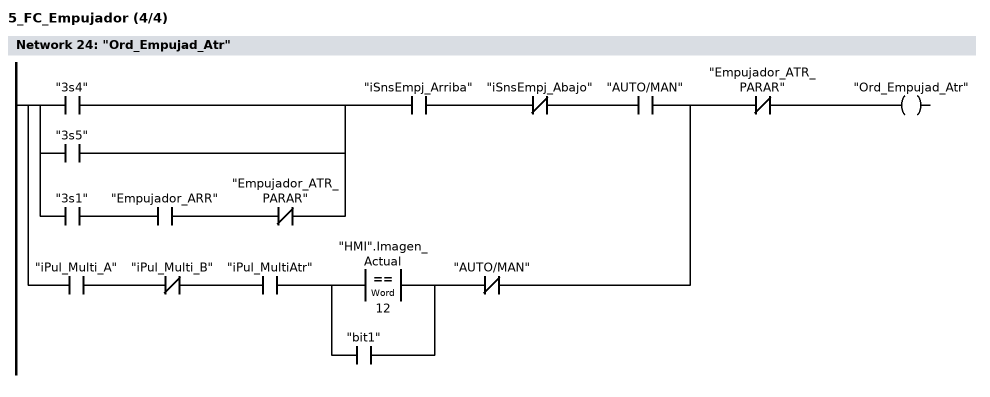
   RUNG wire#powerrail
      Contact( "3s4" )
      wire#w1
      Contact( "iSnsEmpj_Arriba" )
      I_Contact( "iSnsEmpj_Abajo" )
      Contact( "AUTO/MAN" )
      wire#w2
      I_Contact( "Empujador_ATR_PARAR" )
      Coil( "Ord_Empujad_Atr" )
   END_RUNG
   RUNG wire#powerrail
      Contact( "3s5" )
   END_RUNG wire#w1
   RUNG wire#powerrail
      Contact( "3s1" )
      Contact( "Empujador_ARR" )
      I_Contact( "Empujador_ATR_PARAR" )
   END_RUNG wire#w1
   RUNG wire#powerrail
      Contact( "iPul_Multi_A" )
      I_Contact( "iPul_Multi_B" )
      Contact( "iPul_MultiAtr" )
      wire#w3
      { S7_Templates := "SrcType := Word" } EQ_Contact(in1 := "HMI".Imagen_Actual, in2 := 12)
      wire#w4
      I_Contact( "AUTO/MAN" )
   END_RUNG wire#w2
   RUNG wire#w3
      Contact( "bit1" )
   END_RUNG wire#w4
   // the same network as SCL:
   "Ord_Empujad_Atr" := ((("3s4" OR "3s5" OR ("3s1" AND "Empujador_ARR" AND NOT "Empujador_ATR_PARAR")) AND "iSnsEmpj_Arriba" AND NOT "iSnsEmpj_Abajo" AND "AUTO/MAN") OR ("iPul_Multi_A" AND NOT "iPul_Multi_B" AND "iPul_MultiAtr" AND (("HMI".Imagen_Actual = 12) OR "bit1") AND NOT "AUTO/MAN")) AND NOT "Empujador_ATR_PARAR";
END_REGION
END_FUNCTION

FUNCTION "6_FC_Carga_Pallets" : Void   // FC13, LAD
{ S7_Optimized_Access := 'FALSE' }
VERSION : 0.1
BEGIN

REGION Network 1: "Poner_Mordazas"
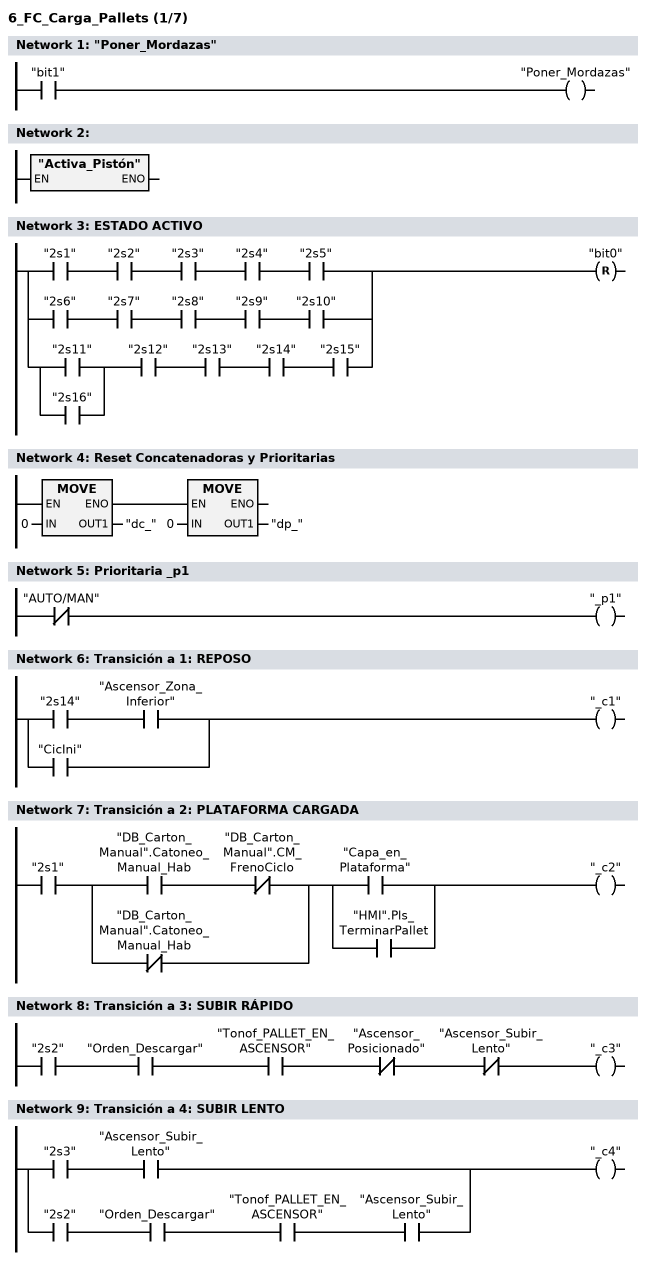
   RUNG wire#powerrail
      Contact( "bit1" )
      Coil( "Poner_Mordazas" )
   END_RUNG
   // the same network as SCL:
   "Poner_Mordazas" := "bit1";
END_REGION

REGION Network 2
   RUNG wire#powerrail
      "Activa_Pistón"()
   END_RUNG
   // the same network as SCL:
   "Activa_Pistón"();
END_REGION

REGION Network 3: ESTADO ACTIVO
   RUNG wire#powerrail
      Contact( "2s1" )
      Contact( "2s2" )
      Contact( "2s3" )
      Contact( "2s4" )
      Contact( "2s5" )
      wire#w1
      R_Coil( "bit0" )
   END_RUNG
   RUNG wire#powerrail
      Contact( "2s6" )
      Contact( "2s7" )
      Contact( "2s8" )
      Contact( "2s9" )
      Contact( "2s10" )
   END_RUNG wire#w1
   RUNG wire#powerrail
      Contact( "2s11" )
      wire#w2
      Contact( "2s12" )
      Contact( "2s13" )
      Contact( "2s14" )
      Contact( "2s15" )
   END_RUNG wire#w1
   RUNG wire#powerrail
      Contact( "2s16" )
   END_RUNG wire#w2
   // the same network as SCL:
   IF ("2s1" AND "2s2" AND "2s3" AND "2s4" AND "2s5") OR ("2s6" AND "2s7" AND "2s8" AND "2s9" AND "2s10") OR (("2s11" OR "2s16") AND "2s12" AND "2s13" AND "2s14" AND "2s15") THEN
       "bit0" := FALSE;
   END_IF;
END_REGION

REGION Network 4: Reset Concatenadoras y Prioritarias
   RUNG wire#powerrail
      { S7_GenerateENO := "TRUE" } Move(in := 0, out1 => "dc_")
      { S7_GenerateENO := "TRUE" } Move(in := 0, out1 => "dp_")
   END_RUNG
   // the same network as SCL:
   // ENO of a box is taken as its EN; it also drops when the box reports an error
   "dc_" := 0;
   "dp_" := 0;
END_REGION

REGION Network 5: Prioritaria _p1
   RUNG wire#powerrail
      I_Contact( "AUTO/MAN" )
      Coil( "_p1" )
   END_RUNG
   // the same network as SCL:
   "_p1" := NOT "AUTO/MAN";
END_REGION

REGION Network 6: Transición a 1: REPOSO
   RUNG wire#powerrail
      Contact( "2s14" )
      Contact( "Ascensor_Zona_Inferior" )
      wire#w1
      Coil( "_c1" )
   END_RUNG
   RUNG wire#powerrail
      Contact( "CicIni" )
   END_RUNG wire#w1
   // the same network as SCL:
   "_c1" := ("2s14" AND "Ascensor_Zona_Inferior") OR "CicIni";
END_REGION

REGION Network 7: Transición a 2: PLATAFORMA CARGADA
   RUNG wire#powerrail
      Contact( "2s1" )
      wire#w1
      Contact( "DB_Carton_Manual".Catoneo_Manual_Hab )
      I_Contact( "DB_Carton_Manual".CM_FrenoCiclo )
      wire#w2
      Contact( "Capa_en_Plataforma" )
      wire#w3
      Coil( "_c2" )
   END_RUNG
   RUNG wire#w1
      I_Contact( "DB_Carton_Manual".Catoneo_Manual_Hab )
   END_RUNG wire#w2
   RUNG wire#w2
      Contact( "HMI".Pls_TerminarPallet )
   END_RUNG wire#w3
   // the same network as SCL:
   "_c2" := "2s1" AND (("DB_Carton_Manual".Catoneo_Manual_Hab AND NOT "DB_Carton_Manual".CM_FrenoCiclo) OR NOT "DB_Carton_Manual".Catoneo_Manual_Hab) AND ("Capa_en_Plataforma" OR "HMI".Pls_TerminarPallet);
END_REGION

REGION Network 8: Transición a 3: SUBIR RÁPIDO
   RUNG wire#powerrail
      Contact( "2s2" )
      Contact( "Orden_Descargar" )
      Contact( "Tonof_PALLET_EN_ASCENSOR" )
      I_Contact( "Ascensor_Posicionado" )
      I_Contact( "Ascensor_Subir_Lento" )
      Coil( "_c3" )
   END_RUNG
   // the same network as SCL:
   "_c3" := "2s2" AND "Orden_Descargar" AND "Tonof_PALLET_EN_ASCENSOR" AND NOT "Ascensor_Posicionado" AND NOT "Ascensor_Subir_Lento";
END_REGION

REGION Network 9: Transición a 4: SUBIR LENTO
   RUNG wire#powerrail
      Contact( "2s3" )
      Contact( "Ascensor_Subir_Lento" )
      wire#w1
      Coil( "_c4" )
   END_RUNG
   RUNG wire#powerrail
      Contact( "2s2" )
      Contact( "Orden_Descargar" )
      Contact( "Tonof_PALLET_EN_ASCENSOR" )
      Contact( "Ascensor_Subir_Lento" )
   END_RUNG wire#w1
   // the same network as SCL:
   "_c4" := ("2s3" AND "Ascensor_Subir_Lento") OR ("2s2" AND "Orden_Descargar" AND "Tonof_PALLET_EN_ASCENSOR" AND "Ascensor_Subir_Lento");
END_REGION

REGION Network 10: Transición a 5: ADELANTAR
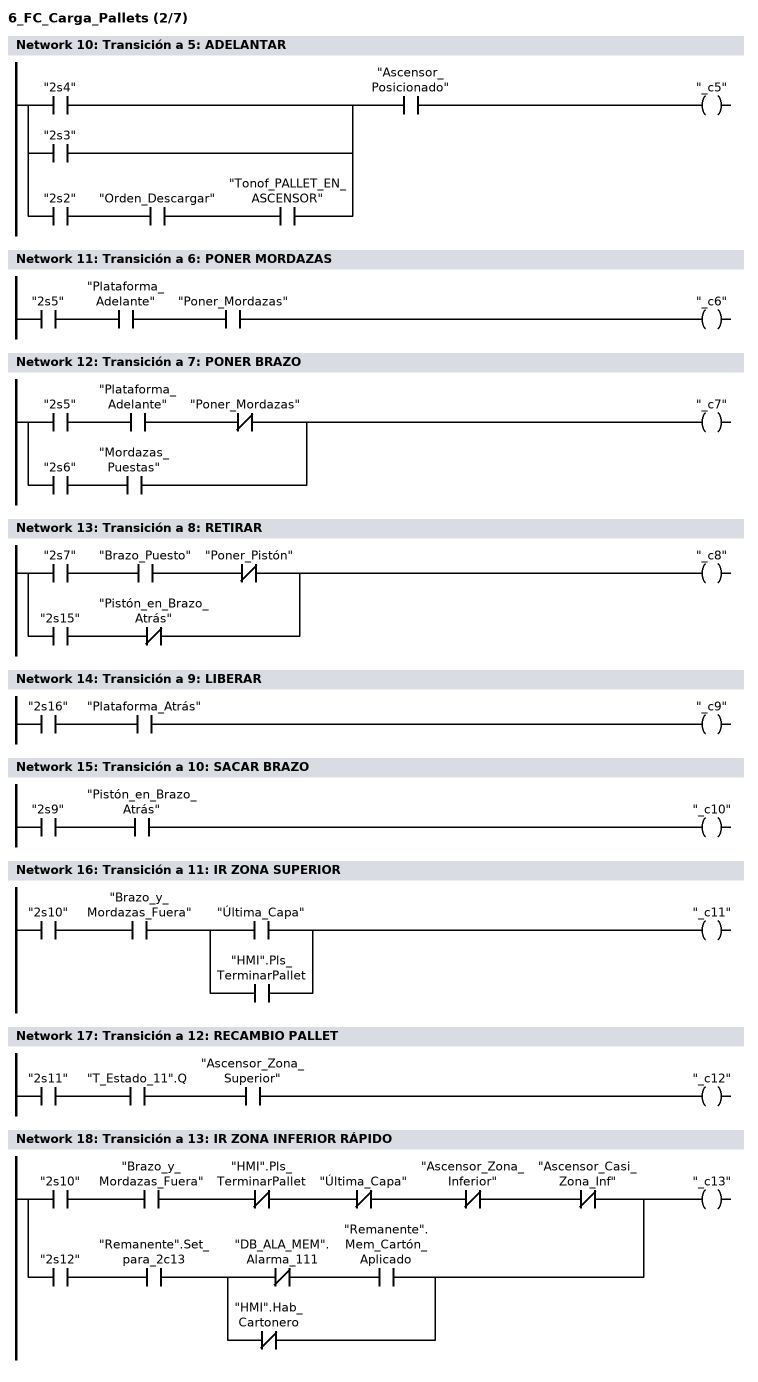
   RUNG wire#powerrail
      Contact( "2s4" )
      wire#w1
      Contact( "Ascensor_Posicionado" )
      Coil( "_c5" )
   END_RUNG
   RUNG wire#powerrail
      Contact( "2s3" )
   END_RUNG wire#w1
   RUNG wire#powerrail
      Contact( "2s2" )
      Contact( "Orden_Descargar" )
      Contact( "Tonof_PALLET_EN_ASCENSOR" )
   END_RUNG wire#w1
   // the same network as SCL:
   "_c5" := ("2s4" OR "2s3" OR ("2s2" AND "Orden_Descargar" AND "Tonof_PALLET_EN_ASCENSOR")) AND "Ascensor_Posicionado";
END_REGION

REGION Network 11: Transición a 6: PONER MORDAZAS
   RUNG wire#powerrail
      Contact( "2s5" )
      Contact( "Plataforma_Adelante" )
      Contact( "Poner_Mordazas" )
      Coil( "_c6" )
   END_RUNG
   // the same network as SCL:
   "_c6" := "2s5" AND "Plataforma_Adelante" AND "Poner_Mordazas";
END_REGION

REGION Network 12: Transición a 7: PONER BRAZO
   RUNG wire#powerrail
      Contact( "2s5" )
      Contact( "Plataforma_Adelante" )
      I_Contact( "Poner_Mordazas" )
      wire#w1
      Coil( "_c7" )
   END_RUNG
   RUNG wire#powerrail
      Contact( "2s6" )
      Contact( "Mordazas_Puestas" )
   END_RUNG wire#w1
   // the same network as SCL:
   "_c7" := ("2s5" AND "Plataforma_Adelante" AND NOT "Poner_Mordazas") OR ("2s6" AND "Mordazas_Puestas");
END_REGION

REGION Network 13: Transición a 8: RETIRAR
   RUNG wire#powerrail
      Contact( "2s7" )
      Contact( "Brazo_Puesto" )
      I_Contact( "Poner_Pistón" )
      wire#w1
      Coil( "_c8" )
   END_RUNG
   RUNG wire#powerrail
      Contact( "2s15" )
      I_Contact( "Pistón_en_Brazo_Atrás" )
   END_RUNG wire#w1
   // the same network as SCL:
   "_c8" := ("2s7" AND "Brazo_Puesto" AND NOT "Poner_Pistón") OR ("2s15" AND NOT "Pistón_en_Brazo_Atrás");
END_REGION

REGION Network 14: Transición a 9: LIBERAR
   RUNG wire#powerrail
      Contact( "2s16" )
      Contact( "Plataforma_Atrás" )
      Coil( "_c9" )
   END_RUNG
   // the same network as SCL:
   "_c9" := "2s16" AND "Plataforma_Atrás";
END_REGION

REGION Network 15: Transición a 10: SACAR BRAZO
   RUNG wire#powerrail
      Contact( "2s9" )
      Contact( "Pistón_en_Brazo_Atrás" )
      Coil( "_c10" )
   END_RUNG
   // the same network as SCL:
   "_c10" := "2s9" AND "Pistón_en_Brazo_Atrás";
END_REGION

REGION Network 16: Transición a 11: IR ZONA SUPERIOR
   RUNG wire#powerrail
      Contact( "2s10" )
      Contact( "Brazo_y_Mordazas_Fuera" )
      wire#w1
      Contact( "Última_Capa" )
      wire#w2
      Coil( "_c11" )
   END_RUNG
   RUNG wire#w1
      Contact( "HMI".Pls_TerminarPallet )
   END_RUNG wire#w2
   // the same network as SCL:
   "_c11" := "2s10" AND "Brazo_y_Mordazas_Fuera" AND ("Última_Capa" OR "HMI".Pls_TerminarPallet);
END_REGION

REGION Network 17: Transición a 12: RECAMBIO PALLET
   RUNG wire#powerrail
      Contact( "2s11" )
      Contact( "T_Estado_11".Q )
      Contact( "Ascensor_Zona_Superior" )
      Coil( "_c12" )
   END_RUNG
   // the same network as SCL:
   "_c12" := "2s11" AND "T_Estado_11".Q AND "Ascensor_Zona_Superior";
END_REGION

REGION Network 18: Transición a 13: IR ZONA INFERIOR RÁPIDO
   RUNG wire#powerrail
      Contact( "2s10" )
      Contact( "Brazo_y_Mordazas_Fuera" )
      I_Contact( "HMI".Pls_TerminarPallet )
      I_Contact( "Última_Capa" )
      I_Contact( "Ascensor_Zona_Inferior" )
      I_Contact( "Ascensor_Casi_Zona_Inf" )
      wire#w1
      Coil( "_c13" )
   END_RUNG
   RUNG wire#powerrail
      Contact( "2s12" )
      Contact( "Remanente".Set_para_2c13 )
      wire#w2
      I_Contact( "DB_ALA_MEM".Alarma_111 )
      Contact( "Remanente".Mem_Cartón_Aplicado )
   END_RUNG wire#w1
   RUNG wire#w2
      I_Contact( "HMI".Hab_Cartonero )
   END_RUNG wire#w1
   // the same network as SCL:
   "_c13" := ("2s10" AND "Brazo_y_Mordazas_Fuera" AND NOT "HMI".Pls_TerminarPallet AND NOT "Última_Capa" AND NOT "Ascensor_Zona_Inferior" AND NOT "Ascensor_Casi_Zona_Inf") OR ("2s12" AND "Remanente".Set_para_2c13 AND ((NOT "DB_ALA_MEM".Alarma_111 AND "Remanente".Mem_Cartón_Aplicado) OR NOT "HMI".Hab_Cartonero));
END_REGION

REGION Network 19: Transición a 14: IR ZONA INFERIOR LENTO
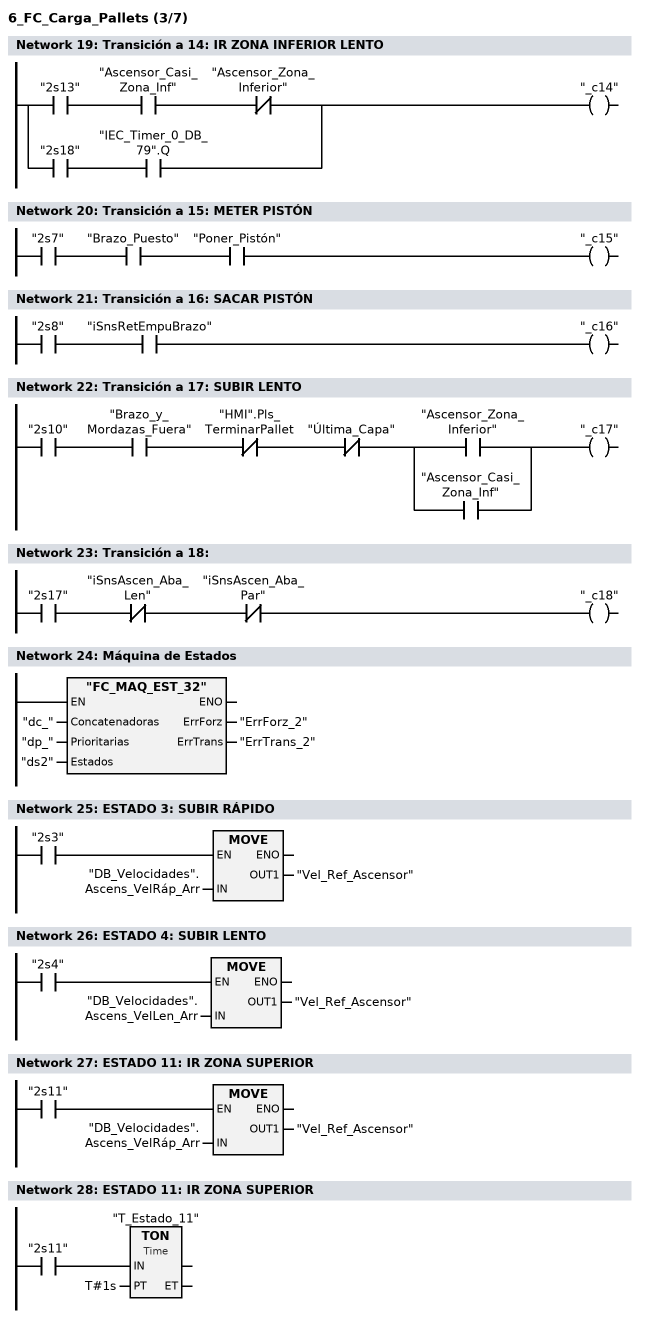
   RUNG wire#powerrail
      Contact( "2s13" )
      Contact( "Ascensor_Casi_Zona_Inf" )
      I_Contact( "Ascensor_Zona_Inferior" )
      wire#w1
      Coil( "_c14" )
   END_RUNG
   RUNG wire#powerrail
      Contact( "2s18" )
      Contact( "IEC_Timer_0_DB_79".Q )
   END_RUNG wire#w1
   // the same network as SCL:
   "_c14" := ("2s13" AND "Ascensor_Casi_Zona_Inf" AND NOT "Ascensor_Zona_Inferior") OR ("2s18" AND "IEC_Timer_0_DB_79".Q);
END_REGION

REGION Network 20: Transición a 15: METER PISTÓN
   RUNG wire#powerrail
      Contact( "2s7" )
      Contact( "Brazo_Puesto" )
      Contact( "Poner_Pistón" )
      Coil( "_c15" )
   END_RUNG
   // the same network as SCL:
   "_c15" := "2s7" AND "Brazo_Puesto" AND "Poner_Pistón";
END_REGION

REGION Network 21: Transición a 16: SACAR PISTÓN
   RUNG wire#powerrail
      Contact( "2s8" )
      Contact( "iSnsRetEmpuBrazo" )
      Coil( "_c16" )
   END_RUNG
   // the same network as SCL:
   "_c16" := "2s8" AND "iSnsRetEmpuBrazo";
END_REGION

REGION Network 22: Transición a 17: SUBIR LENTO
   RUNG wire#powerrail
      Contact( "2s10" )
      Contact( "Brazo_y_Mordazas_Fuera" )
      I_Contact( "HMI".Pls_TerminarPallet )
      I_Contact( "Última_Capa" )
      wire#w1
      Contact( "Ascensor_Zona_Inferior" )
      wire#w2
      Coil( "_c17" )
   END_RUNG
   RUNG wire#w1
      Contact( "Ascensor_Casi_Zona_Inf" )
   END_RUNG wire#w2
   // the same network as SCL:
   "_c17" := "2s10" AND "Brazo_y_Mordazas_Fuera" AND NOT "HMI".Pls_TerminarPallet AND NOT "Última_Capa" AND ("Ascensor_Zona_Inferior" OR "Ascensor_Casi_Zona_Inf");
END_REGION

REGION Network 23: Transición a 18:
   RUNG wire#powerrail
      Contact( "2s17" )
      I_Contact( "iSnsAscen_Aba_Len" )
      I_Contact( "iSnsAscen_Aba_Par" )
      Coil( "_c18" )
   END_RUNG
   // the same network as SCL:
   "_c18" := "2s17" AND NOT "iSnsAscen_Aba_Len" AND NOT "iSnsAscen_Aba_Par";
END_REGION

REGION Network 24: Máquina de Estados
   RUNG wire#powerrail
      "FC_MAQ_EST_32"(Concatenadoras := "dc_", Prioritarias := "dp_", Estados := "ds2", ErrForz => "ErrForz_2", ErrTrans => "ErrTrans_2")
   END_RUNG
   // the same network as SCL:
   "FC_MAQ_EST_32"(Concatenadoras := "dc_",
                   Prioritarias := "dp_",
                   Estados := "ds2",
                   ErrForz => "ErrForz_2",
                   ErrTrans => "ErrTrans_2");
END_REGION

REGION Network 25: ESTADO 3: SUBIR RÁPIDO
   RUNG wire#powerrail
      Contact( "2s3" )
      { S7_GenerateENO := "TRUE" } Move(in := "DB_Velocidades".Ascens_VelRáp_Arr, out1 => "Vel_Ref_Ascensor")
   END_RUNG
   // the same network as SCL:
   IF "2s3" THEN "Vel_Ref_Ascensor" := "DB_Velocidades".Ascens_VelRáp_Arr; END_IF;
END_REGION

REGION Network 26: ESTADO 4: SUBIR LENTO
   RUNG wire#powerrail
      Contact( "2s4" )
      { S7_GenerateENO := "TRUE" } Move(in := "DB_Velocidades".Ascens_VelLen_Arr, out1 => "Vel_Ref_Ascensor")
   END_RUNG
   // the same network as SCL:
   IF "2s4" THEN "Vel_Ref_Ascensor" := "DB_Velocidades".Ascens_VelLen_Arr; END_IF;
END_REGION

REGION Network 27: ESTADO 11: IR ZONA SUPERIOR
   RUNG wire#powerrail
      Contact( "2s11" )
      { S7_GenerateENO := "TRUE" } Move(in := "DB_Velocidades".Ascens_VelRáp_Arr, out1 => "Vel_Ref_Ascensor")
   END_RUNG
   // the same network as SCL:
   IF "2s11" THEN "Vel_Ref_Ascensor" := "DB_Velocidades".Ascens_VelRáp_Arr; END_IF;
END_REGION

REGION Network 28: ESTADO 11: IR ZONA SUPERIOR
   "T_Estado_11".TON(in := "2s11", pt := T#1s);
END_REGION

REGION Network 29: ESTADO 12: RECAMBIO PALLET
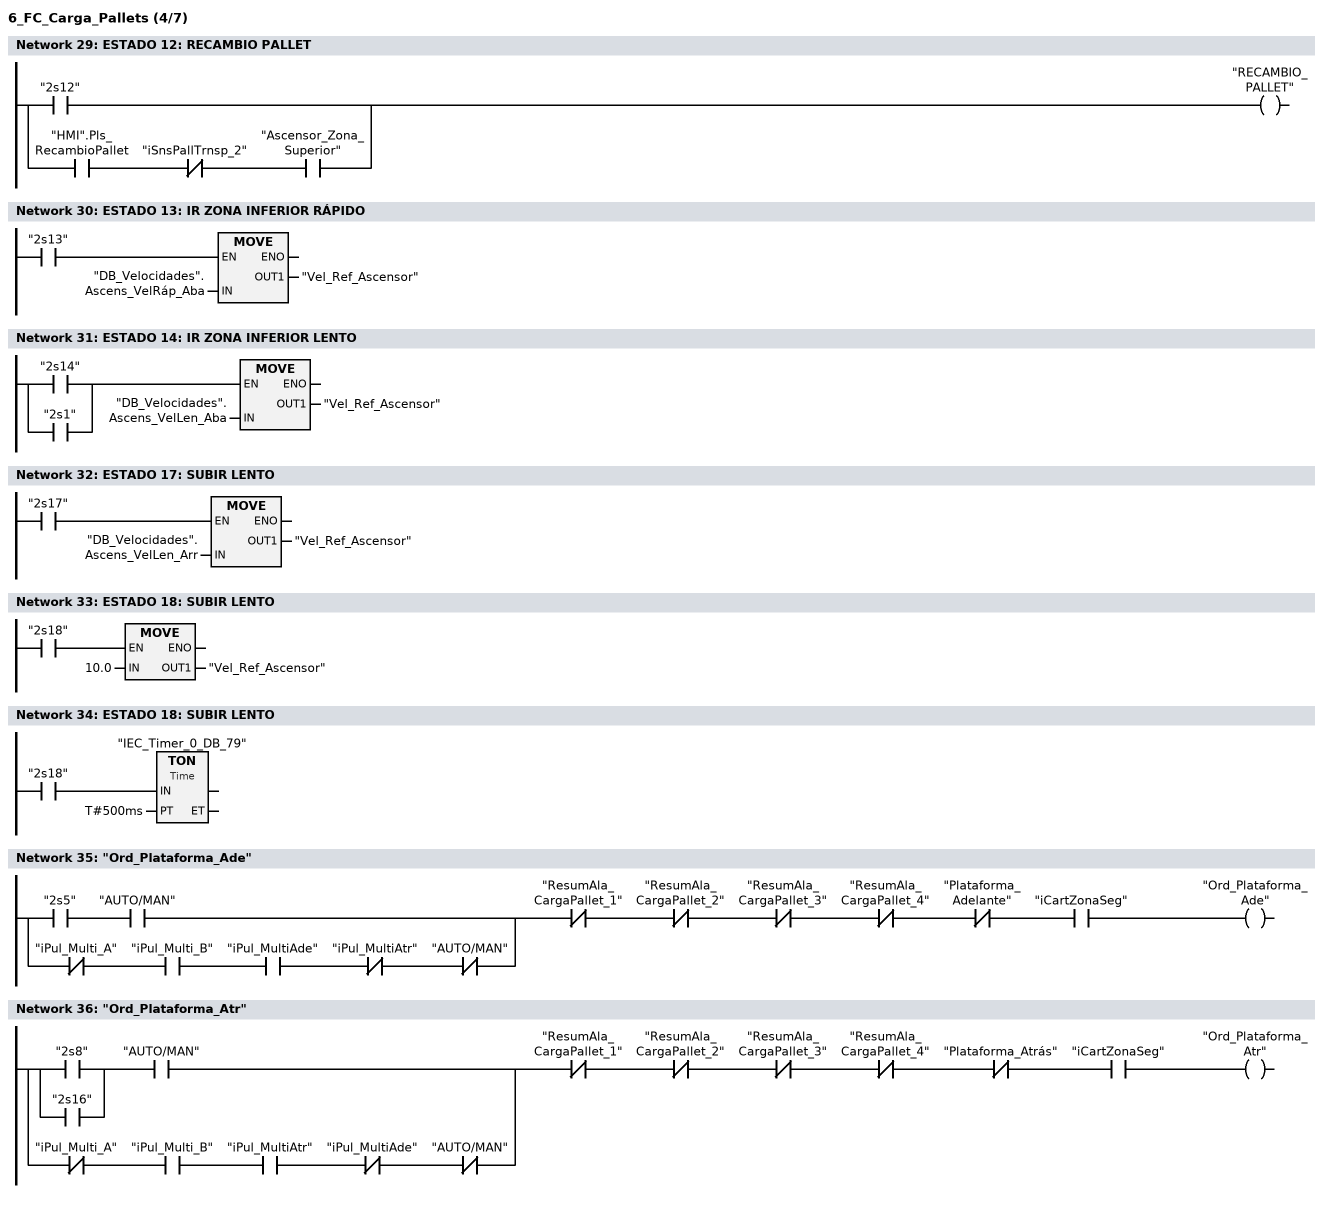
   RUNG wire#powerrail
      Contact( "2s12" )
      wire#w1
      Coil( "RECAMBIO_PALLET" )
   END_RUNG
   RUNG wire#powerrail
      Contact( "HMI".Pls_RecambioPallet )
      I_Contact( "iSnsPallTrnsp_2" )
      Contact( "Ascensor_Zona_Superior" )
   END_RUNG wire#w1
   // the same network as SCL:
   "RECAMBIO_PALLET" := "2s12" OR ("HMI".Pls_RecambioPallet AND NOT "iSnsPallTrnsp_2" AND "Ascensor_Zona_Superior");
END_REGION

REGION Network 30: ESTADO 13: IR ZONA INFERIOR RÁPIDO
   RUNG wire#powerrail
      Contact( "2s13" )
      { S7_GenerateENO := "TRUE" } Move(in := "DB_Velocidades".Ascens_VelRáp_Aba, out1 => "Vel_Ref_Ascensor")
   END_RUNG
   // the same network as SCL:
   IF "2s13" THEN "Vel_Ref_Ascensor" := "DB_Velocidades".Ascens_VelRáp_Aba; END_IF;
END_REGION

REGION Network 31: ESTADO 14: IR ZONA INFERIOR LENTO
   RUNG wire#powerrail
      Contact( "2s14" )
      wire#w1
      { S7_GenerateENO := "TRUE" } Move(in := "DB_Velocidades".Ascens_VelLen_Aba, out1 => "Vel_Ref_Ascensor")
   END_RUNG
   RUNG wire#powerrail
      Contact( "2s1" )
   END_RUNG wire#w1
   // the same network as SCL:
   IF "2s14" OR "2s1" THEN "Vel_Ref_Ascensor" := "DB_Velocidades".Ascens_VelLen_Aba; END_IF;
END_REGION

REGION Network 32: ESTADO 17: SUBIR LENTO
   RUNG wire#powerrail
      Contact( "2s17" )
      { S7_GenerateENO := "TRUE" } Move(in := "DB_Velocidades".Ascens_VelLen_Arr, out1 => "Vel_Ref_Ascensor")
   END_RUNG
   // the same network as SCL:
   IF "2s17" THEN "Vel_Ref_Ascensor" := "DB_Velocidades".Ascens_VelLen_Arr; END_IF;
END_REGION

REGION Network 33: ESTADO 18: SUBIR LENTO
   RUNG wire#powerrail
      Contact( "2s18" )
      { S7_GenerateENO := "TRUE" } Move(in := 10.0, out1 => "Vel_Ref_Ascensor")
   END_RUNG
   // the same network as SCL:
   IF "2s18" THEN "Vel_Ref_Ascensor" := 10.0; END_IF;
END_REGION

REGION Network 34: ESTADO 18: SUBIR LENTO
   "IEC_Timer_0_DB_79".TON(in := "2s18", pt := T#500ms);
END_REGION

REGION Network 35: "Ord_Plataforma_Ade"
   RUNG wire#powerrail
      Contact( "2s5" )
      Contact( "AUTO/MAN" )
      wire#w1
      I_Contact( "ResumAla_CargaPallet_1" )
      I_Contact( "ResumAla_CargaPallet_2" )
      I_Contact( "ResumAla_CargaPallet_3" )
      I_Contact( "ResumAla_CargaPallet_4" )
      I_Contact( "Plataforma_Adelante" )
      Contact( "iCartZonaSeg" )
      Coil( "Ord_Plataforma_Ade" )
   END_RUNG
   RUNG wire#powerrail
      I_Contact( "iPul_Multi_A" )
      Contact( "iPul_Multi_B" )
      Contact( "iPul_MultiAde" )
      I_Contact( "iPul_MultiAtr" )
      I_Contact( "AUTO/MAN" )
   END_RUNG wire#w1
   // the same network as SCL:
   "Ord_Plataforma_Ade" := (("2s5" AND "AUTO/MAN") OR (NOT "iPul_Multi_A" AND "iPul_Multi_B" AND "iPul_MultiAde" AND NOT "iPul_MultiAtr" AND NOT "AUTO/MAN")) AND NOT "ResumAla_CargaPallet_1" AND NOT "ResumAla_CargaPallet_2" AND NOT "ResumAla_CargaPallet_3" AND NOT "ResumAla_CargaPallet_4" AND NOT "Plataforma_Adelante" AND "iCartZonaSeg";
END_REGION

REGION Network 36: "Ord_Plataforma_Atr"
   RUNG wire#powerrail
      Contact( "2s8" )
      wire#w1
      Contact( "AUTO/MAN" )
      wire#w2
      I_Contact( "ResumAla_CargaPallet_1" )
      I_Contact( "ResumAla_CargaPallet_2" )
      I_Contact( "ResumAla_CargaPallet_3" )
      I_Contact( "ResumAla_CargaPallet_4" )
      I_Contact( "Plataforma_Atrás" )
      Contact( "iCartZonaSeg" )
      Coil( "Ord_Plataforma_Atr" )
   END_RUNG
   RUNG wire#powerrail
      Contact( "2s16" )
   END_RUNG wire#w1
   RUNG wire#powerrail
      I_Contact( "iPul_Multi_A" )
      Contact( "iPul_Multi_B" )
      Contact( "iPul_MultiAtr" )
      I_Contact( "iPul_MultiAde" )
      I_Contact( "AUTO/MAN" )
   END_RUNG wire#w2
   // the same network as SCL:
   "Ord_Plataforma_Atr" := ((("2s8" OR "2s16") AND "AUTO/MAN") OR (NOT "iPul_Multi_A" AND "iPul_Multi_B" AND "iPul_MultiAtr" AND NOT "iPul_MultiAde" AND NOT "AUTO/MAN")) AND NOT "ResumAla_CargaPallet_1" AND NOT "ResumAla_CargaPallet_2" AND NOT "ResumAla_CargaPallet_3" AND NOT "ResumAla_CargaPallet_4" AND NOT "Plataforma_Atrás" AND "iCartZonaSeg";
END_REGION

REGION Network 37: "Ord_Ascensor_Subir"
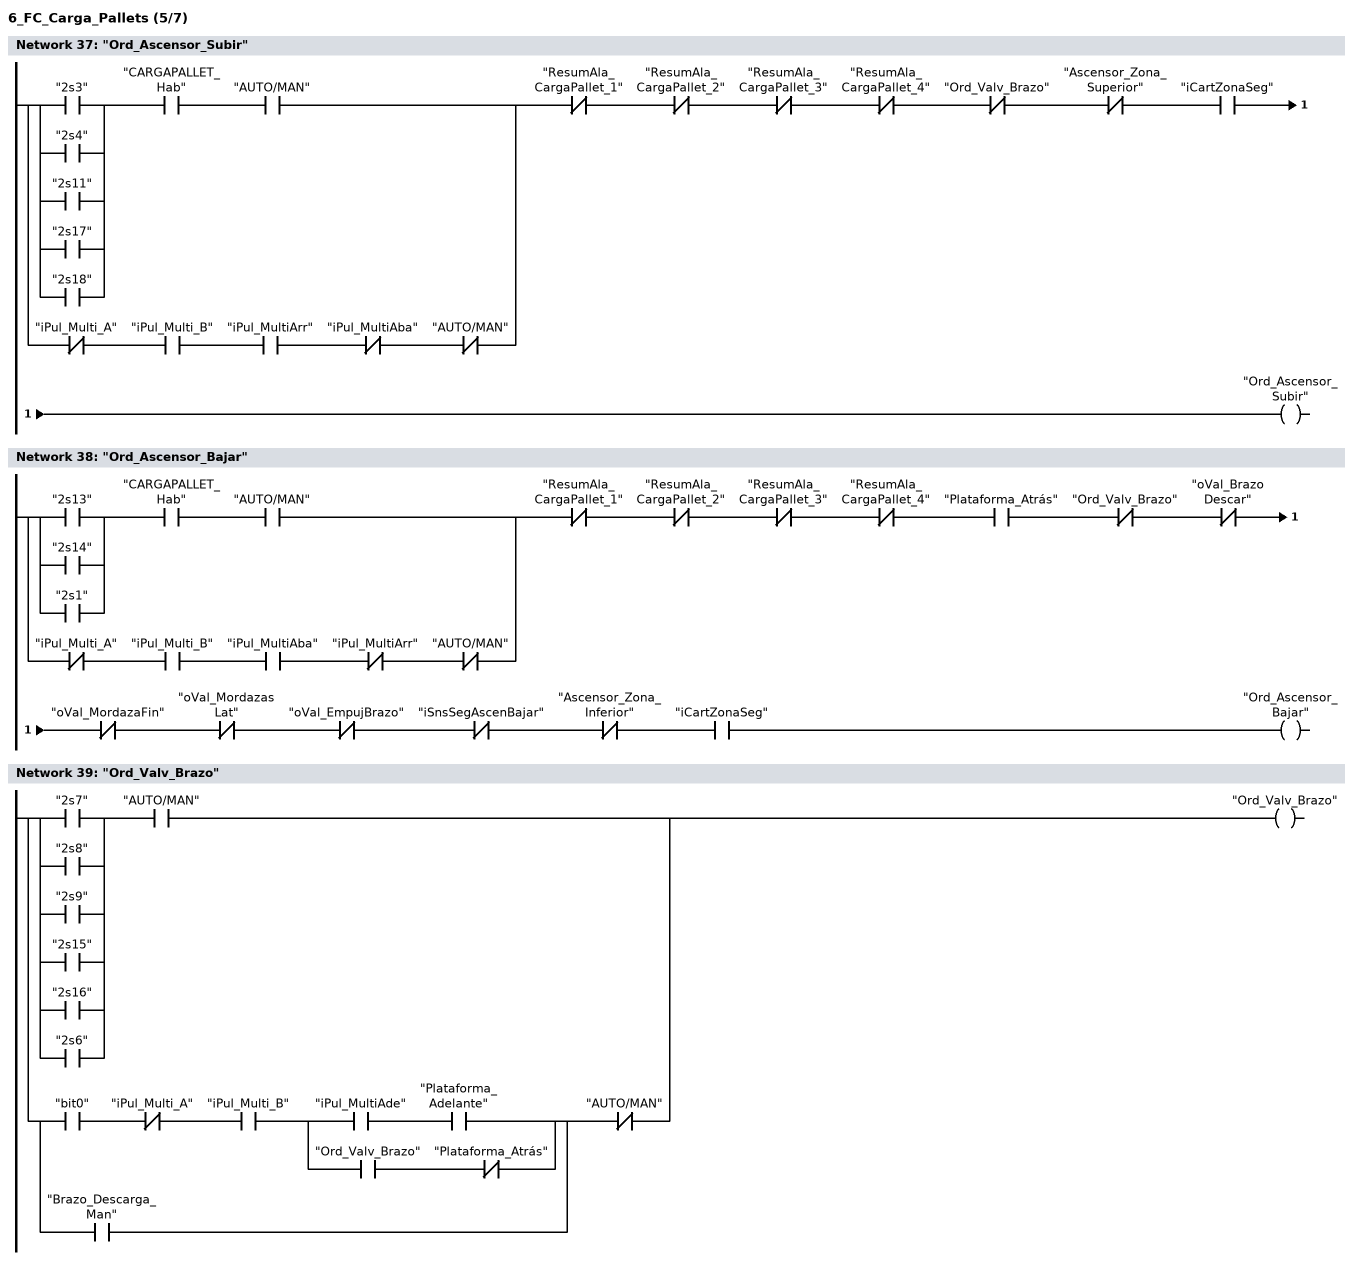
   RUNG wire#powerrail
      Contact( "2s3" )
      wire#w1
      Contact( "CARGAPALLET_Hab" )
      Contact( "AUTO/MAN" )
      wire#w2
      I_Contact( "ResumAla_CargaPallet_1" )
      I_Contact( "ResumAla_CargaPallet_2" )
      I_Contact( "ResumAla_CargaPallet_3" )
      I_Contact( "ResumAla_CargaPallet_4" )
      I_Contact( "Ord_Valv_Brazo" )
      I_Contact( "Ascensor_Zona_Superior" )
      Contact( "iCartZonaSeg" )
      Coil( "Ord_Ascensor_Subir" )
   END_RUNG
   RUNG wire#powerrail
      Contact( "2s4" )
   END_RUNG wire#w1
   RUNG wire#powerrail
      Contact( "2s11" )
   END_RUNG wire#w1
   RUNG wire#powerrail
      Contact( "2s17" )
   END_RUNG wire#w1
   RUNG wire#powerrail
      Contact( "2s18" )
   END_RUNG wire#w1
   RUNG wire#powerrail
      I_Contact( "iPul_Multi_A" )
      Contact( "iPul_Multi_B" )
      Contact( "iPul_MultiArr" )
      I_Contact( "iPul_MultiAba" )
      I_Contact( "AUTO/MAN" )
   END_RUNG wire#w2
   // the same network as SCL:
   "Ord_Ascensor_Subir" := ((("2s3" OR "2s4" OR "2s11" OR "2s17" OR "2s18") AND "CARGAPALLET_Hab" AND "AUTO/MAN") OR (NOT "iPul_Multi_A" AND "iPul_Multi_B" AND "iPul_MultiArr" AND NOT "iPul_MultiAba" AND NOT "AUTO/MAN")) AND NOT "ResumAla_CargaPallet_1" AND NOT "ResumAla_CargaPallet_2" AND NOT "ResumAla_CargaPallet_3" AND NOT "ResumAla_CargaPallet_4" AND NOT "Ord_Valv_Brazo" AND NOT "Ascensor_Zona_Superior" AND "iCartZonaSeg";
END_REGION

REGION Network 38: "Ord_Ascensor_Bajar"
   RUNG wire#powerrail
      Contact( "2s13" )
      wire#w1
      Contact( "CARGAPALLET_Hab" )
      Contact( "AUTO/MAN" )
      wire#w2
      I_Contact( "ResumAla_CargaPallet_1" )
      I_Contact( "ResumAla_CargaPallet_2" )
      I_Contact( "ResumAla_CargaPallet_3" )
      I_Contact( "ResumAla_CargaPallet_4" )
      Contact( "Plataforma_Atrás" )
      I_Contact( "Ord_Valv_Brazo" )
      I_Contact( "oVal_BrazoDescar" )
      I_Contact( "oVal_MordazaFin" )
      I_Contact( "oVal_MordazasLat" )
      I_Contact( "oVal_EmpujBrazo" )
      I_Contact( "iSnsSegAscenBajar" )
      I_Contact( "Ascensor_Zona_Inferior" )
      Contact( "iCartZonaSeg" )
      Coil( "Ord_Ascensor_Bajar" )
   END_RUNG
   RUNG wire#powerrail
      Contact( "2s14" )
   END_RUNG wire#w1
   RUNG wire#powerrail
      Contact( "2s1" )
   END_RUNG wire#w1
   RUNG wire#powerrail
      I_Contact( "iPul_Multi_A" )
      Contact( "iPul_Multi_B" )
      Contact( "iPul_MultiAba" )
      I_Contact( "iPul_MultiArr" )
      I_Contact( "AUTO/MAN" )
   END_RUNG wire#w2
   // the same network as SCL:
   "Ord_Ascensor_Bajar" := ((("2s13" OR "2s14" OR "2s1") AND "CARGAPALLET_Hab" AND "AUTO/MAN") OR (NOT "iPul_Multi_A" AND "iPul_Multi_B" AND "iPul_MultiAba" AND NOT "iPul_MultiArr" AND NOT "AUTO/MAN")) AND NOT "ResumAla_CargaPallet_1" AND NOT "ResumAla_CargaPallet_2" AND NOT "ResumAla_CargaPallet_3" AND NOT "ResumAla_CargaPallet_4" AND "Plataforma_Atrás" AND NOT "Ord_Valv_Brazo" AND NOT "oVal_BrazoDescar" AND NOT "oVal_MordazaFin" AND NOT "oVal_MordazasLat" AND NOT "oVal_EmpujBrazo" AND NOT "iSnsSegAscenBajar" AND NOT "Ascensor_Zona_Inferior" AND "iCartZonaSeg";
END_REGION

REGION Network 39: "Ord_Valv_Brazo"
   RUNG wire#powerrail
      Contact( "2s7" )
      wire#w1
      Contact( "AUTO/MAN" )
      wire#w2
      Coil( "Ord_Valv_Brazo" )
   END_RUNG
   RUNG wire#powerrail
      Contact( "2s8" )
   END_RUNG wire#w1
   RUNG wire#powerrail
      Contact( "2s9" )
   END_RUNG wire#w1
   RUNG wire#powerrail
      Contact( "2s15" )
   END_RUNG wire#w1
   RUNG wire#powerrail
      Contact( "2s16" )
   END_RUNG wire#w1
   RUNG wire#powerrail
      Contact( "2s6" )
   END_RUNG wire#w1
   RUNG wire#powerrail
      Contact( "bit0" )
      I_Contact( "iPul_Multi_A" )
      Contact( "iPul_Multi_B" )
      wire#w3
      Contact( "iPul_MultiAde" )
      Contact( "Plataforma_Adelante" )
      wire#w4
      I_Contact( "AUTO/MAN" )
   END_RUNG wire#w2
   RUNG wire#w3
      Contact( "Ord_Valv_Brazo" )
      I_Contact( "Plataforma_Atrás" )
   END_RUNG wire#w4
   RUNG wire#powerrail
      Contact( "Brazo_Descarga_Man" )
   END_RUNG wire#w4
   // the same network as SCL:
   "Ord_Valv_Brazo" := (("2s7" OR "2s8" OR "2s9" OR "2s15" OR "2s16" OR "2s6") AND "AUTO/MAN") OR ((("bit0" AND NOT "iPul_Multi_A" AND "iPul_Multi_B" AND (("iPul_MultiAde" AND "Plataforma_Adelante") OR ("Ord_Valv_Brazo" AND NOT "Plataforma_Atrás"))) OR "Brazo_Descarga_Man") AND NOT "AUTO/MAN");
END_REGION

REGION Network 40: "Ord_Valv_Pistón_Brazo"
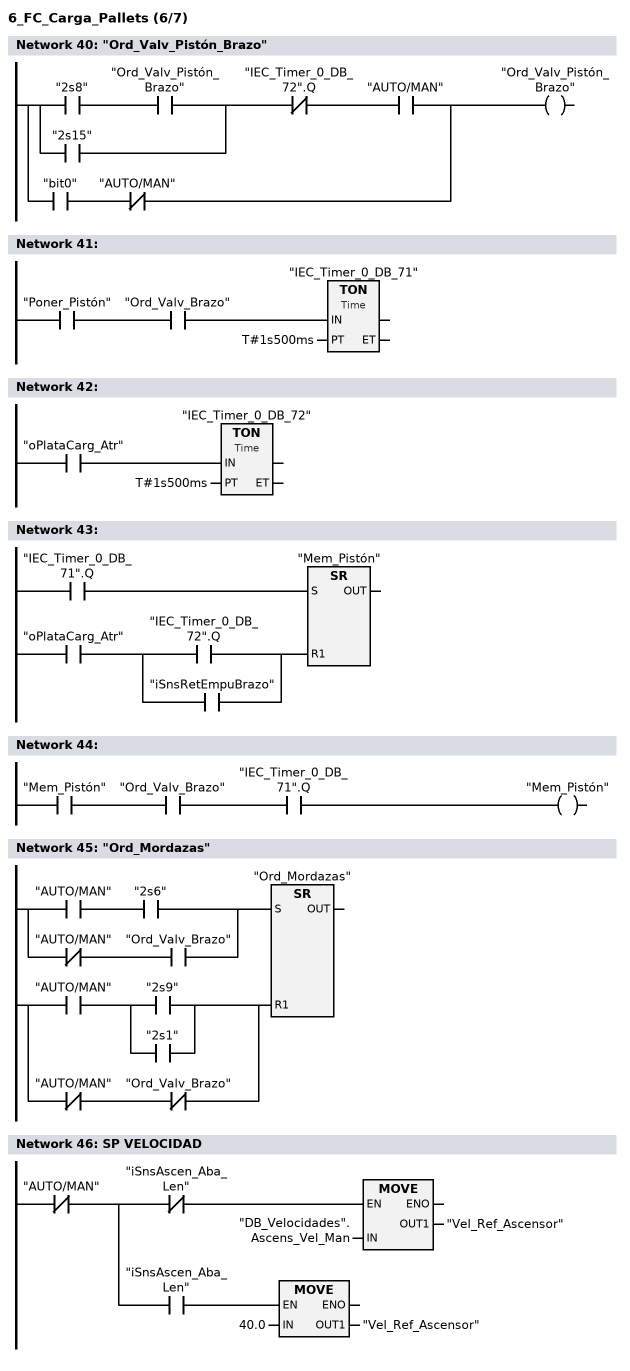
   RUNG wire#powerrail
      Contact( "2s8" )
      Contact( "Ord_Valv_Pistón_Brazo" )
      wire#w1
      I_Contact( "IEC_Timer_0_DB_72".Q )
      Contact( "AUTO/MAN" )
      wire#w2
      Coil( "Ord_Valv_Pistón_Brazo" )
   END_RUNG
   RUNG wire#powerrail
      Contact( "2s15" )
   END_RUNG wire#w1
   RUNG wire#powerrail
      Contact( "bit0" )
      I_Contact( "AUTO/MAN" )
   END_RUNG wire#w2
   // the same network as SCL:
   "Ord_Valv_Pistón_Brazo" := ((("2s8" AND "Ord_Valv_Pistón_Brazo") OR "2s15") AND NOT "IEC_Timer_0_DB_72".Q AND "AUTO/MAN") OR ("bit0" AND NOT "AUTO/MAN");
END_REGION

REGION Network 41
   "IEC_Timer_0_DB_71".TON(in := "Poner_Pistón" AND "Ord_Valv_Brazo", pt := T#1s500ms);
END_REGION

REGION Network 42
   "IEC_Timer_0_DB_72".TON(in := "oPlataCarg_Atr", pt := T#1s500ms);
END_REGION

REGION Network 43
   RUNG wire#powerrail
      Contact( "IEC_Timer_0_DB_71".Q )
      S_SR(operand := "Mem_Pistón", r1 := wire#w2)
   END_RUNG
   RUNG wire#powerrail
      Contact( "oPlataCarg_Atr" )
      wire#w1
      Contact( "IEC_Timer_0_DB_72".Q )
   END_RUNG wire#w2
   RUNG wire#w1
      Contact( "iSnsRetEmpuBrazo" )
   END_RUNG wire#w2
   // the same network as SCL:
   IF "IEC_Timer_0_DB_71".Q THEN
       "Mem_Pistón" := TRUE;   // SR flip-flop
   END_IF;
   IF "oPlataCarg_Atr" AND ("IEC_Timer_0_DB_72".Q OR "iSnsRetEmpuBrazo") THEN "Mem_Pistón" := FALSE; END_IF;
END_REGION

REGION Network 44
   RUNG wire#powerrail
      Contact( "Mem_Pistón" )
      Contact( "Ord_Valv_Brazo" )
      Contact( "IEC_Timer_0_DB_71".Q )
      Coil( "Mem_Pistón" )
   END_RUNG
   // the same network as SCL:
   "Mem_Pistón" := "Mem_Pistón" AND "Ord_Valv_Brazo" AND "IEC_Timer_0_DB_71".Q;
END_REGION

REGION Network 45: "Ord_Mordazas"
   RUNG wire#powerrail
      Contact( "AUTO/MAN" )
      Contact( "2s6" )
      wire#w1
      S_SR(operand := "Ord_Mordazas", r1 := wire#w3)
   END_RUNG
   RUNG wire#powerrail
      I_Contact( "AUTO/MAN" )
      Contact( "Ord_Valv_Brazo" )
   END_RUNG wire#w1
   RUNG wire#powerrail
      Contact( "AUTO/MAN" )
      wire#w2
      Contact( "2s9" )
   END_RUNG wire#w3
   RUNG wire#w2
      Contact( "2s1" )
   END_RUNG wire#w3
   RUNG wire#powerrail
      I_Contact( "AUTO/MAN" )
      I_Contact( "Ord_Valv_Brazo" )
   END_RUNG wire#w3
   // the same network as SCL:
   IF ("AUTO/MAN" AND "2s6") OR (NOT "AUTO/MAN" AND "Ord_Valv_Brazo") THEN
       "Ord_Mordazas" := TRUE;   // SR flip-flop
   END_IF;
   IF ("AUTO/MAN" AND ("2s9" OR "2s1")) OR (NOT "AUTO/MAN" AND NOT "Ord_Valv_Brazo") THEN
       "Ord_Mordazas" := FALSE;
   END_IF;
END_REGION

REGION Network 46: SP VELOCIDAD
   RUNG wire#powerrail
      I_Contact( "AUTO/MAN" )
      wire#w1
      I_Contact( "iSnsAscen_Aba_Len" )
      { S7_GenerateENO := "TRUE" } Move(in := "DB_Velocidades".Ascens_Vel_Man, out1 => "Vel_Ref_Ascensor")
   END_RUNG
   RUNG wire#w1
      Contact( "iSnsAscen_Aba_Len" )
      { S7_GenerateENO := "TRUE" } Move(in := 40.0, out1 => "Vel_Ref_Ascensor")
   END_RUNG
   // the same network as SCL:
   IF NOT "AUTO/MAN" AND NOT "iSnsAscen_Aba_Len" THEN
       "Vel_Ref_Ascensor" := "DB_Velocidades".Ascens_Vel_Man;
   END_IF;
   IF NOT "AUTO/MAN" AND "iSnsAscen_Aba_Len" THEN "Vel_Ref_Ascensor" := 40.0; END_IF;
END_REGION

REGION Network 47: "TON_AcumPalet"
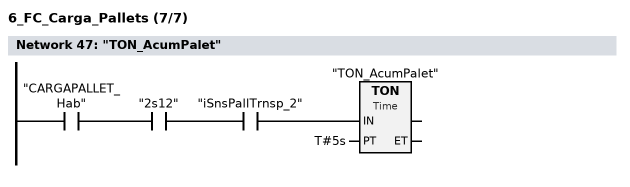
   "TON_AcumPalet".TON(IN := "CARGAPALLET_Hab" AND "2s12" AND "iSnsPallTrnsp_2", PT := T#5s);
END_REGION
END_FUNCTION

FUNCTION "7_FC_Transp_Pallets" : Void   // FC14, LAD
{ S7_Optimized_Access := 'FALSE' }
VERSION : 0.1
BEGIN

REGION Network 1: Pallet_Transporte1_a_Transporte2